// TIA Portal project "Robotino" (V18)

(* hardware
DEVICE "S7-1500/ET200MP-Station_1"  S7-1500 station
   slot 0: "Profilschiene_0"  Rack  6ES7 590-1***0-0AA0
   slot 1: "PLC_1"  CPU 1516-3 PN/DP  6ES7 516-3AP03-0AB0  V3.0
      slot 3: "CPU-Display_1"  6ES7591-1BA00-0AA0
      slot 32768: "PROFINET-Schnittstelle_1"  X1
      slot 33024: "PROFINET-Schnittstelle_2"  X2
      slot 33280: "DP-Schnittstelle_1"  X3
      slot 34817: "Virtual CP interface port_1"  Virtual CP interface port  Virtual CP interface port
   slot 2: "DI 32x24VDC HF_1"  DI 32x24VDC HF  6ES7 521-1BL00-0AB0  V2.2
   slot 3: "DQ 32x24VDC/0.5A HF_1"  DQ 32x24VDC/0.5A HF  6ES7 522-1BL01-0AB0  V1.1
   slot 4: "AI 8xU/I/RTD/TC ST_1"  AI 8xU/I/RTD/TC ST  6ES7 531-7KF00-0AB0  V2.2
   slot 5: "AQ 4xU/I ST_1"  AQ 4xU/I ST  6ES7 532-5HD00-0AB0  V2.2
DEVICE "ROBOTINO_HMI"  MTP700 Unified Comfort
   slot 0: "ROBOTINO_HMI"  MTP700 Unified Comfort  6AV2 128-3GB06-0AXx  18.0.0.2
   slot 1: "HMI_RT_1"  MTP700 Unified Comfort  6AV2 128-3GB06-0AXx  18.0.0.2
   slot 5: "ROBOTINO_HMI.IE_CP_1"  PROFINET Interface  18.0.0.2
      slot 1: "PROFINET Schnittstelle_1"  PROFINET Interface
         slot 1: "Port_1"  Port
         slot 2: "Port_2"  Port
   slot 6: "ROBOTINO_HMI.IE_CP_2"  PROFINET Interface  18.0.0.2
      slot 1: "PROFINET Schnittstelle_GBit"  PROFINET Interface
         slot 1: "Port_1"  Port
*)

// ===== PLC "PLC_1"  CPU 1516-3 PN/DP =====

DATA_BLOCK "OPCUA"   // DB1
{ S7_Optimized_Access := 'TRUE' }
VERSION : 0.1
   VAR
      Test_bool : Bool;
      Test_int : Int;
      Test_String : String;
      Test_array_bool : Array[0..1] of Bool;
      Test_array_int : Array[0..1] of Int;
   END_VAR
BEGIN
END_DATA_BLOCK

DATA_BLOCK "ROBOTINO"   // DB2
{ S7_Optimized_Access := 'TRUE' }
VERSION : 0.1
   VAR
      Bumper : Bool;
      Distance_Sensors : Array[1..9] of Real;
      Digital_Inputs : Array[1..8] of Bool;
      Analog_Inputs : Array[1..8] of Real;
      Motor4 : Int;   // Belt
      Motor4_Current : Real;
      Digital_Outputs : Array[1..8] of Bool;
      Digital_Outputs_Status : Array[1..8] of Bool;
      Relay : Array[1..2] of Bool;
      Relay_Status : Array[1..2] of Bool;
      Odometry : Array[0..6] of Real;
      Omnidrive : Array[0..2] of Real;
      Bat_Voltage : Real;
      Charging_State : String;
      Charging_Current : Real;
      Controller_Info : Array[0..1] of String;
      Image_Version : String;
      Factory_Status : Array[0..3] of Bool;
      Position_ID : Int;
      Start_GoToPos : Bool;
      GoToPos_Completed : Bool;
      Robotino_Position : Int;   // actual defined position of robotino. =0 If robotino is not on a defined position
      DockTo_Completed : Bool;   // =1 if robotino is docked
      Start_DockTo : Bool;
      Stop_DockTo : Bool;
   END_VAR
BEGIN
   // Digital_Inputs[3] : Vision Sensor Package Present
   // Digital_Inputs[4] : IR Station Ready (false connected)
   // Digital_Inputs[5] : Reset Button
   // Digital_Outputs[3] : lamp tower red
   // Digital_Outputs[4] : lamp tower yellow
   // Digital_Outputs[5] : lamp tower green
   // Digital_Outputs[6] : light reset button
   // Digital_Outputs[1] : IR Robotino Ready
   // Digital_Outputs_Status[1] : IR Robotino Ready
   // Digital_Outputs_Status[3] : lamp tower red
   // Digital_Outputs_Status[4] : lamp tower yellow
   // Digital_Outputs_Status[5] : lamp tower green
   // Digital_Outputs_Status[6] : light reset button
   // Relay_Status[1] : Enable analog sensors
   // Odometry[0] : x /m
   // Odometry[1] : y /m
   // Odometry[2] : rot /rad
   // Odometry[3] : vx
   // Odometry[4] : vy
   // Odometry[5] : omega
   // Odometry[6] : sequence number
   // Omnidrive[0] : vx
   // Omnidrive[1] : vy
   // Omnidrive[2] : omega
   // Relay[1] : Enable analog sensors
   // Analog_Inputs[1] : Distance Left (not scaled)
   // Analog_Inputs[2] : Distance Center (not scaled)
   // Analog_Inputs[3] : Distance Right (not scaled)
   // Controller_Info[1] : Software version
   // Controller_Info[0] : Hardware version
   // Factory_Status[0] : Idle
   // Factory_Status[1] : Busy
   // Factory_Status[2] : Error
   // Factory_Status[3] : Started
   // Digital_Inputs[1] : Emergncy Button
END_DATA_BLOCK

DATA_BLOCK "GoTo_DB"   // DB3
{ S7_Optimized_Access := 'TRUE' }
VERSION : 0.1
// stored: InstanceOfName GoTo
"GoTo"
BEGIN
END_DATA_BLOCK

DATA_BLOCK "DockTo_DB"   // DB5
{ S7_Optimized_Access := 'TRUE' }
VERSION : 0.1
// stored: InstanceOfName DockTo
"DockTo"
BEGIN
END_DATA_BLOCK

DATA_BLOCK "Robotino_Control"   // DB6
{ S7_Optimized_Access := 'TRUE' }
VERSION : 0.1
   VAR
      Start_GoTo : Bool;
      Start_DockTo : Bool;
      Ready_DockTo : Bool;
      Stop_DockTo : Bool;
      Conveyor : Int;
      PosId : Int;
   END_VAR
BEGIN
END_DATA_BLOCK

// folder: System blocks/Program resources

DATA_BLOCK "IEC_Timer_0_DB"   // DB4
{ S7_Optimized_Access := 'TRUE' }
AUTHOR : Simatic
FAMILY : IEC
NAME : IEC_TMR
VERSION : 1.0
// stored: InstanceOfName IEC_TIMER
"IEC_TIMER"
BEGIN
END_DATA_BLOCK

DATA_BLOCK "IEC_Timer_0_DB_1"   // DB8
{ S7_Optimized_Access := 'TRUE' }
AUTHOR : Simatic
FAMILY : IEC
NAME : IEC_TMR
VERSION : 1.0
// stored: InstanceOfName IEC_TIMER
"IEC_TIMER"
BEGIN
END_DATA_BLOCK

// folder: (top level)

FUNCTION_BLOCK "GoTo"   // FB1, FBD
{ S7_Optimized_Access := 'TRUE' }
VERSION : 0.1
   VAR_INPUT
      Idle : Bool;
      Busy : Bool;
      Error : Bool;
      Started : Bool;
      Pos : Int;
      Start : Bool;
   END_VAR
   VAR_OUTPUT
      GoTo_Completed : Bool;
      GoTo_Start : Bool;
      GoTo_PosId : Int;
      actual_PosId : Int;
   END_VAR
   VAR_TEMP
      process_completed : Bool;
      busy_negedge : Bool;
      idle_posedge : Bool;
      process_started : Bool;
      completed_p_edge : Bool;
   END_VAR
   VAR_TEMP   // added for the SCL form of the ladder/FBD networks
      _w1 : Bool;
   END_VAR
BEGIN

REGION Network 1
   // Anzahl definierter Positionen in Factory ggf. anpassen
   // 
   // Sinnhaftigkeit von TOF und Zeit prüfen
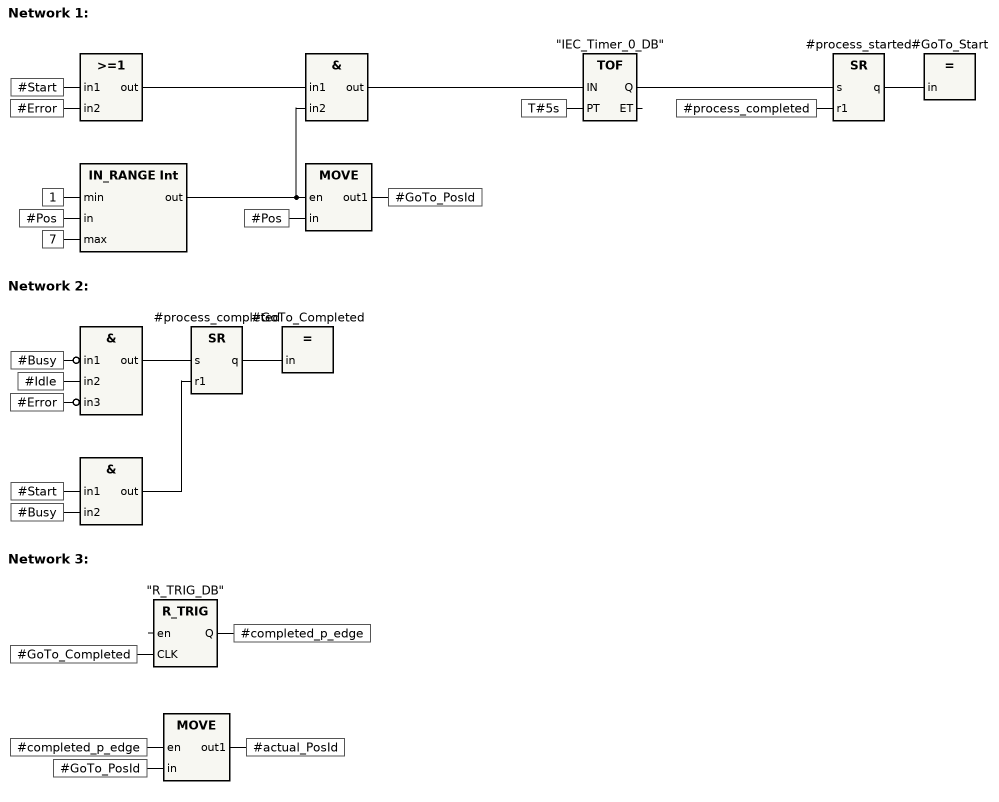
   #_w1 := (1 <= #Pos) AND (#Pos <= 7);
   "IEC_Timer_0_DB".TOF(IN := (#Start OR #Error) AND #_w1, PT := T#5s);
   IF "IEC_Timer_0_DB".Q THEN
       #process_started := TRUE;   // SR flip-flop
   END_IF;
   IF #process_completed THEN #process_started := FALSE; END_IF;
   #GoTo_Start := #process_started;
   IF #_w1 THEN #GoTo_PosId := #Pos; END_IF;
END_REGION

REGION Network 2
   // Startbefehl nach GoToCompleted zurückssetzen
   IF NOT #Busy AND #Idle AND NOT #Error THEN
       #process_completed := TRUE;   // SR flip-flop
   END_IF;
   IF #Start AND #Busy THEN #process_completed := FALSE; END_IF;
   #GoTo_Completed := #process_completed;
END_REGION

REGION Network 3
   // Registrierung der aktuellen Position
   // nur p edge als enable nehemen
   "R_TRIG_DB"(CLK := #GoTo_Completed, Q => #completed_p_edge);   // R_TRIG
   IF #completed_p_edge THEN #actual_PosId := #GoTo_PosId; END_IF;
END_REGION
END_FUNCTION_BLOCK

FUNCTION_BLOCK "DockTo"   // FB2, GRAPH_PLUS
{ S7_Optimized_Access := 'TRUE' }
VERSION : 0.1
   VAR_INPUT
      OFF_SQ : Bool := false;
      INIT_SQ : Bool := false;
      ACK_EF : Bool := false;
      S_PREV : Bool := false;
      S_NEXT : Bool := false;
      SW_AUTO : Bool := false;
      SW_TAP : Bool := false;
      SW_TOP : Bool := false;
      SW_MAN : Bool := false;
      S_SEL : Int := 0;
      S_ON : Bool := false;
      S_OFF : Bool := false;
      T_PUSH : Bool := false;
      idle : Bool;
      busy : Bool;
      error_factory : Bool;
      robotino_position : Int;
      distance_left : Real;
      distance_center : Real;
      distance_right : Real;
   END_VAR
   VAR_OUTPUT
      S_NO : Int := 0;
      S_MORE : Bool := false;
      S_ACTIVE : Bool := false;
      ERR_FLT : Bool := false;
      AUTO_ON : Bool := false;
      TAP_ON : Bool := false;
      TOP_ON : Bool := false;
      MAN_ON : Bool := false;
      docking_completed : Bool;
      docking_started : Bool;
      vx : Real;
      vy : Real;
      omega : Real;
      relay_analogsensors : Bool;
   END_VAR
   VAR
      HMI_INFO : Array[0..8] of UInt;
      IF_PAR : G7_IfParPlus_V6;
      RT_DATA : G7_RTDataPlus_V6;
      Trans1 : G7_TransitionPlus_V6;
      Trans2 : G7_TransitionPlus_V6;
      Trans3 : G7_TransitionPlus_V6;
      Trans4 : G7_TransitionPlus_V6;
      Trans5 : G7_TransitionPlus_V6;
      Trans6 : G7_TransitionPlus_V6;
      Trans7 : G7_TransitionPlus_V6;
      Trans8 : G7_TransitionPlus_V6;   // Transitionsstruktur
      Trans9 : G7_TransitionPlus_V6;   // Transitionsstruktur
      Trans10 : G7_TransitionPlus_V6;   // Transitionsstruktur
      Trans11 : G7_TransitionPlus_V6;   // Transitionsstruktur
      Trans13 : G7_TransitionPlus_V6;   // Transitionsstruktur
      Trans14 : G7_TransitionPlus_V6;   // Transitionsstruktur
      Trans18 : G7_TransitionPlus_V6;   // Transitionsstruktur
      Step1 : G7_StepPlus_V6;
      Step2 : G7_StepPlus_V6;
      Step3 : G7_StepPlus_V6;
      Step4 : G7_StepPlus_V6;
      Step5 : G7_StepPlus_V6;
      Step6 : G7_StepPlus_V6;
      Step7 : G7_StepPlus_V6;   // Schrittstruktur
      Step8 : G7_StepPlus_V6;   // Schrittstruktur
      Step9 : G7_StepPlus_V6;   // Schrittstruktur
      Step11 : G7_StepPlus_V6;   // Schrittstruktur
      Step13 : G7_StepPlus_V6;   // Schrittstruktur
      Step14 : G7_StepPlus_V6;   // Schrittstruktur
      SINI : Array[0..1] of USInt;
      LSTT : Array[0..13] of USInt;
      ATAJ : Array[0..13] of USInt;
      ATAB : Array[0..13] of USInt;
      PSTT : Array[0..13] of USInt;
      NSTT : Array[0..13] of USInt;
      ASSJ : Array[0..11] of USInt;
      ASSB : Array[0..11] of USInt;
      PTTS : Array[0..11] of USInt;
      NTTS : Array[0..11] of USInt;
      SW_SQTS : Array[0..11] of USInt;
      SWITCH : Array[0..6] of USInt;
      TVX : Array[0..5] of USInt;
      TTX : Array[0..5] of USInt;
      TSX : Array[0..1] of USInt;
      S00X : Array[0..1] of USInt;
      SOFFX : Array[0..1] of USInt;
      SONX : Array[0..1] of USInt;
      SAX : Array[0..1] of USInt;
      SERRX : Array[0..12] of USInt;
      SMX : Array[0..12] of USInt;
      S0X : Array[0..12] of USInt;
      S1X : Array[0..12] of USInt;
      IL_ALARM_INST : Diag_Alarm;
      SUP_ALARM_INST : Diag_Alarm;
      STEP_TIME_ALARM_INST : Diag_Alarm;
      IEC_TIMER_INST : IEC_TIMER;
      TRANSACTION_FLAG : Bool := false;
   END_VAR
   VAR CONSTANT
      threshold_x : Real := 1.5;
      threshold_y : Real := 1.4;
   END_VAR
   // SINI[0] := 2;
   // LSTT[0] := 255;
   // ATAJ[1] := 1;
   // ATAB[1] := 1;
   // PSTT[1] := 1;
   // NSTT[0] := 3;
   // ASSJ[1] := 1;
   // ASSB[1] := 1;
   // PTTS[0] := 255;
   // NTTS[1] := 1;
   // TVX[0] := 16#1;
   // TTX[0] := 16#1;
   // TSX[0] := 16#1;
   // S00X[0] := 16#1;
   // SOFFX[0] := 16#1;
   // SONX[0] := 16#1;
   // SAX[0] := 16#1;
   // SERRX[0] := 16#1;
   // SMX[0] := 16#1;
   // S0X[0] := 16#1;
   // S1X[0] := 16#1;
   // LSTT[1] := 255;
   // ATAJ[2] := 2;
   // ATAB[2] := 2;
   // PSTT[2] := 2;
   // NSTT[1] := 6;
   // ASSJ[2] := 2;
   // ASSB[2] := 2;
   // PTTS[2] := 9;
   // NTTS[2] := 2;
   // LSTT[3] := 255;
   // LSTT[4] := 255;
   // LSTT[5] := 255;
   // LSTT[6] := 255;
   // ATAJ[3] := 3;
   // ATAJ[4] := 4;
   // ATAJ[5] := 5;
   // ATAJ[6] := 6;
   // ATAB[3] := 4;
   // ATAB[4] := 3;
   // ATAB[5] := 5;
   // ATAB[6] := 6;
   // PSTT[3] := 3;
   // PSTT[4] := 3;
   // PSTT[5] := 5;
   // PSTT[6] := 4;
   // NSTT[3] := 5;
   // NSTT[4] := 4;
   // NSTT[5] := 1;
   // NSTT[6] := 10;
   // ASSJ[3] := 3;
   // ASSJ[4] := 4;
   // ASSJ[5] := 5;
   // ASSB[3] := 3;
   // ASSB[4] := 4;
   // ASSB[5] := 5;
   // PTTS[1] := 5;
   // PTTS[4] := 4;
   // PTTS[5] := 3;
   // NTTS[3] := 3;
   // NTTS[4] := 6;
   // NTTS[5] := 5;
   // SW_SQTS[1] := 1;
   // SW_SQTS[2] := 2;
   // SW_SQTS[4] := 3;
   // SW_SQTS[5] := 1;
   // LSTT[7] := 255;
   // ATAJ[7] := 7;
   // ATAB[7] := 8;
   // PSTT[7] := 9;
   // NSTT[7] := 7;
   // ASSJ[6] := 6;
   // ASSB[6] := 6;
   // PTTS[6] := 1;
   // NTTS[6] := 11;
   // SW_SQTS[6] := 1;
   // LSTT[8] := 255;
   // LSTT[9] := 255;
   // LSTT[10] := 255;
   // ATAJ[8] := 8;
   // ATAJ[9] := 10;
   // ATAJ[10] := 9;
   // ATAB[8] := 7;
   // ATAB[9] := 9;
   // ATAB[10] := 10;
   // PSTT[8] := 9;
   // PSTT[9] := 7;
   // PSTT[10] := 8;
   // NSTT[8] := 8;
   // NSTT[9] := 2;
   // NSTT[10] := 2;
   // ASSJ[7] := 7;
   // ASSJ[8] := 8;
   // ASSB[7] := 7;
   // ASSB[8] := 8;
   // PTTS[7] := 7;
   // PTTS[8] := 8;
   // NTTS[7] := 9;
   // NTTS[8] := 10;
   // SW_SQTS[7] := 4;
   // SW_SQTS[8] := 5;
   // LSTT[11] := 255;
   // LSTT[12] := 255;
   // LSTT[13] := 255;
   // ATAJ[11] := 13;
   // ATAJ[12] := 12;
   // ATAJ[13] := 11;
   // ATAB[11] := 11;
   // ATAB[12] := 12;
   // ATAB[13] := 13;
   // PSTT[11] := 6;
   // PSTT[12] := 10;
   // PSTT[13] := 11;
   // NSTT[11] := 9;
   // NSTT[12] := 11;
   // NSTT[13] := 9;
   // ASSJ[9] := 9;
   // ASSJ[10] := 10;
   // ASSJ[11] := 11;
   // ASSB[9] := 9;
   // ASSB[10] := 10;
   // ASSB[11] := 11;
   // PTTS[9] := 11;
   // PTTS[10] := 6;
   // PTTS[11] := 12;
   // NTTS[9] := 7;
   // NTTS[10] := 12;
   // NTTS[11] := 13;
   // SW_SQTS[9] := 6;
   // SW_SQTS[10] := 3;
   // SW_SQTS[11] := 3;
BEGIN
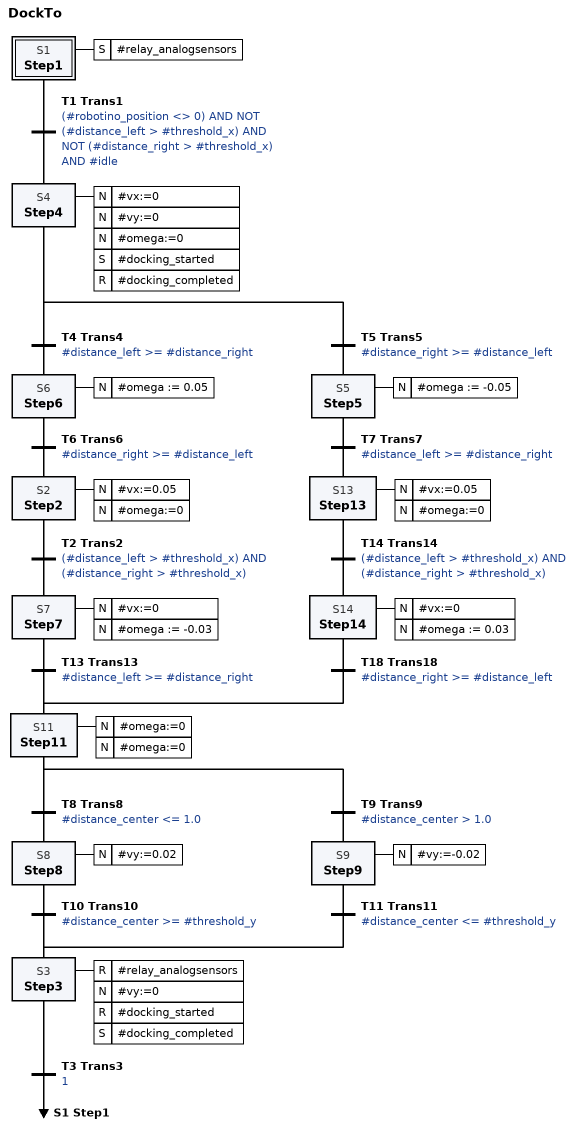
   // sequencer 1
   INITIAL_STEP Step1:   // S1, max time T#10S, warning time T#7S
              S    #relay_analogsensors
   END_STEP
   TRANSITION Trans1 FROM Step1 TO Step4   // T1
      := (#robotino_position <> 0) AND NOT (#distance_left > #threshold_x) AND NOT (#distance_right > #threshold_x) AND #idle;
   END_TRANSITION
   STEP Step2:   // S2, max time T#10S, warning time T#7S
              N    #vx:=0.05
              N    #omega:=0
   END_STEP
   TRANSITION Trans2 FROM Step2 TO Step7   // T2
      := (#distance_left > #threshold_x) AND (#distance_right > #threshold_x);
   END_TRANSITION
   STEP Step3:   // S3, max time T#10S, warning time T#7S
              R    #relay_analogsensors
              N    #vy:=0
              R    #docking_started
              S    #docking_completed
   END_STEP
   TRANSITION Trans3 FROM Step3 TO Step1   // T3, jump
      := 1;
   END_TRANSITION
   STEP Step4:   // S4, max time T#10S, warning time T#7S
              N    #vx:=0
              N    #vy:=0
              N    #omega:=0
              S    #docking_started
              R    #docking_completed
   END_STEP
   TRANSITION Trans4 FROM Step4 TO Step6   // T4
      := #distance_left >= #distance_right;
   END_TRANSITION
   TRANSITION Trans5 FROM Step4 TO Step5   // T5
      := #distance_right >= #distance_left;
   END_TRANSITION
   STEP Step5:   // S5, max time T#10S, warning time T#7S
              N    #omega := -0.05
   END_STEP
   TRANSITION Trans7 FROM Step5 TO Step13   // T7
      := #distance_left >= #distance_right;
   END_TRANSITION
   STEP Step6:   // S6, max time T#10S, warning time T#7S
              N    #omega := 0.05
   END_STEP
   TRANSITION Trans6 FROM Step6 TO Step2   // T6
      := #distance_right >= #distance_left;
   END_TRANSITION
   STEP Step7:   // S7, max time T#10S, warning time T#7S
              N    #vx:=0
              N    #omega := -0.03
   END_STEP
   TRANSITION Trans13 FROM Step7 TO Step11   // T13
      := #distance_left >= #distance_right;
   END_TRANSITION
   STEP Step8:   // S8, max time T#10S, warning time T#7S
              N    #vy:=0.02
   END_STEP
   TRANSITION Trans10 FROM Step8 TO Step3   // T10
      := #distance_center >= #threshold_y;
   END_TRANSITION
   STEP Step9:   // S9, max time T#10S, warning time T#7S
              N    #vy:=-0.02
   END_STEP
   TRANSITION Trans11 FROM Step9 TO Step3   // T11
      := #distance_center <= #threshold_y;
   END_TRANSITION
   STEP Step11:   // S11, max time T#10S, warning time T#7S
              N    #omega:=0
              N    #omega:=0
   END_STEP
   TRANSITION Trans8 FROM Step11 TO Step8   // T8
      := #distance_center <= 1.0;
   END_TRANSITION
   TRANSITION Trans9 FROM Step11 TO Step9   // T9
      := #distance_center > 1.0;
   END_TRANSITION
   STEP Step13:   // S13, max time T#10S, warning time T#7S
              N    #vx:=0.05
              N    #omega:=0
   END_STEP
   TRANSITION Trans14 FROM Step13 TO Step14   // T14
      := (#distance_left > #threshold_x) AND (#distance_right > #threshold_x);
   END_TRANSITION
   STEP Step14:   // S14, max time T#10S, warning time T#7S
              N    #vx:=0
              N    #omega := 0.03
   END_STEP
   TRANSITION Trans18 FROM Step14 TO Step11   // T18
      := #distance_right >= #distance_left;
   END_TRANSITION
END_FUNCTION_BLOCK

ORGANIZATION_BLOCK "Main"   // OB1, FBD, ProgramCycle
{ S7_Optimized_Access := 'TRUE' }
VERSION : 0.1
   VAR_INPUT
      Initial_Call : Bool;
      Remanence : Bool;
   END_VAR
BEGIN

REGION Network 1: HMI
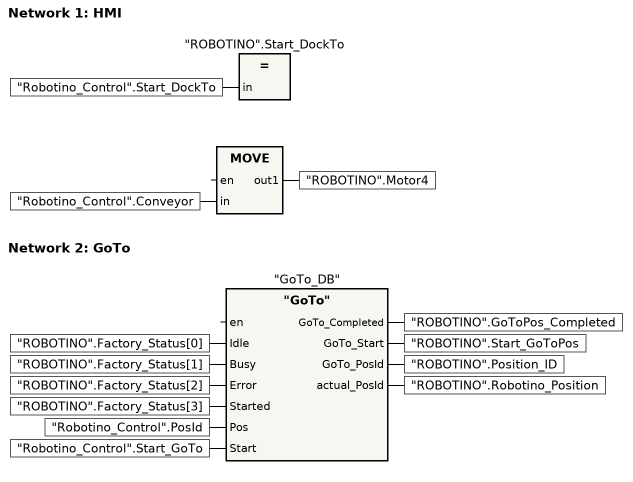
   "ROBOTINO".Start_DockTo := "Robotino_Control".Start_DockTo;
   "ROBOTINO".Motor4 := "Robotino_Control".Conveyor;
END_REGION

REGION Network 2: GoTo
   "GoTo_DB"(Idle := "ROBOTINO".Factory_Status[0],   // "GoTo"
             Busy := "ROBOTINO".Factory_Status[1],
             Error := "ROBOTINO".Factory_Status[2],
             Started := "ROBOTINO".Factory_Status[3],
             Pos := "Robotino_Control".PosId,
             Start := "Robotino_Control".Start_GoTo,
             GoTo_Completed => "ROBOTINO".GoToPos_Completed,
             GoTo_Start => "ROBOTINO".Start_GoToPos,
             GoTo_PosId => "ROBOTINO".Position_ID,
             actual_PosId => "ROBOTINO".Robotino_Position);
END_REGION

REGION Network 3: DockTo
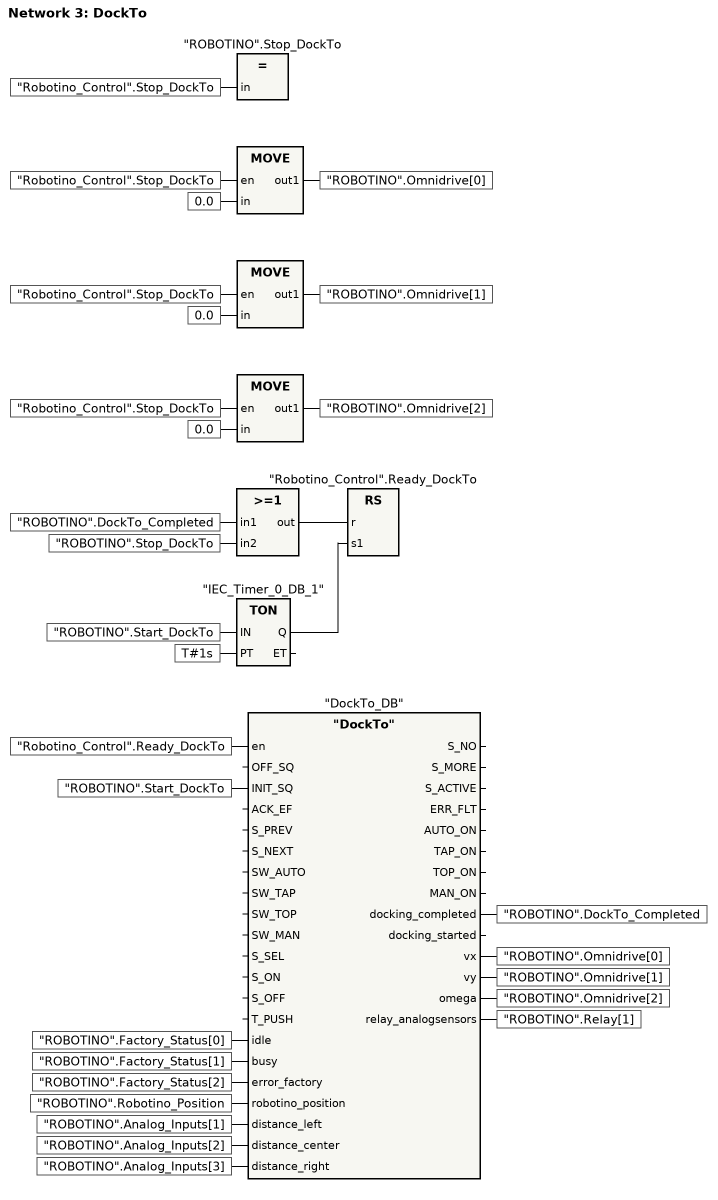
   "ROBOTINO".Stop_DockTo := "Robotino_Control".Stop_DockTo;
   IF "Robotino_Control".Stop_DockTo THEN
       "ROBOTINO".Omnidrive[0] := 0.0;
       "ROBOTINO".Omnidrive[1] := 0.0;
       "ROBOTINO".Omnidrive[2] := 0.0;
   END_IF;
   "IEC_Timer_0_DB_1".TON(IN := "ROBOTINO".Start_DockTo, PT := T#1s);
   IF "ROBOTINO".DockTo_Completed OR "ROBOTINO".Stop_DockTo THEN
       "Robotino_Control".Ready_DockTo := FALSE;   // RS flip-flop
   END_IF;
   IF "IEC_Timer_0_DB_1".Q THEN "Robotino_Control".Ready_DockTo := TRUE; END_IF;
   IF "Robotino_Control".Ready_DockTo THEN
       "DockTo_DB"(INIT_SQ := "ROBOTINO".Start_DockTo,   // "DockTo"
                   idle := "ROBOTINO".Factory_Status[0],
                   busy := "ROBOTINO".Factory_Status[1],
                   error_factory := "ROBOTINO".Factory_Status[2],
                   robotino_position := "ROBOTINO".Robotino_Position,
                   distance_left := "ROBOTINO".Analog_Inputs[1],
                   distance_center := "ROBOTINO".Analog_Inputs[2],
                   distance_right := "ROBOTINO".Analog_Inputs[3],
                   docking_completed => "ROBOTINO".DockTo_Completed,
                   vx => "ROBOTINO".Omnidrive[0],
                   vy => "ROBOTINO".Omnidrive[1],
                   omega => "ROBOTINO".Omnidrive[2],
                   relay_analogsensors => "ROBOTINO".Relay[1]);
   END_IF;
END_REGION
END_ORGANIZATION_BLOCK

(* ===== HMI "HMI_RT_1" =====
connection "HMI_Verbindung_1": ETHERNET, ILRT_S7_1500_OMS

HMI tags "Standard-Variablentabelle"
   "Robotino_Control_Start_GoTo" : Bool = PLC Robotino_Control.Start_GoTo, T100ms
   "Robotino_Control_Start_DockTo" : Bool = PLC Robotino_Control.Start_DockTo, T100ms
   "Robotino_Control_Stop_DockTo" : Bool = PLC Robotino_Control.Stop_DockTo, T100ms
   "Robotino_Control_Conveyor" : Int = PLC Robotino_Control.Conveyor, T100ms
   "Robotino_Control_PosId" : Int = PLC Robotino_Control.PosId, T100ms
   "ROBOTINO_Digital_Inputs{1}" : Bool = PLC ROBOTINO.Digital_Inputs[1] AT %DB1.DBW0, T100ms
   "ROBOTINO_Digital_Outputs_Status{3}" : Bool = PLC ROBOTINO.Digital_Outputs_Status[3], T100ms
   "ROBOTINO_Digital_Outputs_Status{4}" : Bool = PLC ROBOTINO.Digital_Outputs_Status[4], T100ms
   "ROBOTINO_Digital_Outputs_Status{5}" : Bool = PLC ROBOTINO.Digital_Outputs_Status[5], T100ms

text list "SystemTextList_ConfigErrorAlarmTextLibrary_1": 1 'NameService Konfigurationsfehler: Implizites Löschen. Subelement-Instanz @6%s@ muss explizit gelöscht werden.'; 2 'NameService Konfigurationsfehler: Implizites Löschen. Alias/Format/Unit-Instanz @6%s@ muss explizit gelöscht werden.'

text list "SystemTextList_ConfigErrorAlarmTextLibrary_2": 1 'EvDpManager::cleanupDeletedDatapoint - alert handler config is deleted implicitly for deleted datapoint, @3%s@'; 2 'EvDpManager::cleanupDeletedDatapoint - alert handler config is deleted implicitly but still has overrides, @3%s@'; 3 'EvDpManager::cleanupDeletedDatapoint - default value config is deleted implicitly for deleted datapoint, @3%s@'; 4 'EvDpManager::cleanupDeletedDatapoint - default value config is deleted implicitly but still has overrides, @3%s@'; 5 'EvDpManager::cleanupDeletedDatapoint - initial value config is deleted implicitly for deleted datapoint, @3%s@'; 6 'EvDpManager::cleanupDeletedDatapoint - initial value config is deleted implicitly but still has overrides, @3%s@'; 7 'EvDpManager::cleanupDeletedDatapoint - distribution config is deleted implicitly for deleted datapoint, @3%s@'; 8 'EvDpManager::cleanupDeletedDatapoint - distribution config is deleted implicitly but still has overrides, @3%s@'; 9 'EvDpManager::cleanupDeletedDatapoint - rangeCheck config is deleted implicitly for deleted datapoint, @3%s@'; 10 'EvDpManager::cleanupDeletedDatapoint - rangeCheck config is deleted implicitly but still has overrides, @3%s@'

text list "SystemTextList_ConfigErrorAlarmTextLibrary_3": 1 'Der konfigurierte Datenpunkttyp wurde gelöscht. Ein konfigurierter Typ ist aber noch für den Knotentyp definiert: @3%s@.'; 2 'Der konfigurierter Datenpunkt-Knotentyp wurde im Datenpunkttyp gelöscht. Ein konfigurierter Typ ist aber noch für das Element definiert: @3%s@.'

text list "SystemTextList_ConfigErrorAlarmTextLibrary_4": 2 'Zyklen: @6%s@ existiert nicht'; 3 'Alarme: @6%s@ existiert bereits'; 4 'Variablen: Adresse @6%s@ wurde abgelehnt'; 1 'Verbindungen: @6%s@ existiert nicht'; 5 'Variablen: Erfassungsart @6%s@ wird nicht unterstützt.'; 6 'Zyklen: @6%s@ wurde gelöscht aber zugehörige Variablen existieren.'; 7 'Verbindungen: @6%s@ wurde gelöscht aber zugehörige Variablen existieren.'; 8 'Variablen: Variable @6%s@ wurde abgelehnt.'; 9 'Variablen: Variable @6%s@ hat einen ungültigen Wert.'; 0 'Verbindungen: Verbindung zu @6%s@ konnte nicht hergestellt werden.'; 65638 'Verbindungen: Verbindung zu @6%s@ konnte nicht hergestellt werden.'; 65639 'Verbindungen: @6%s@ getrennt.'; 65640 'Verbindungen: Verbindung zum HMI-Gerät @6%s@ getrennt.'; 65641 'Verbindungen: Verbindung zur PLC @6%s@ getrennt.'; 65541 'Verbindungen: Zeitüberschreitung beim Aufbau der Verbindung zu @6%s@.'; 65542 'Verbindungen: @6%s@ gestört.'; 65543 'Verbindungen: Verbindung zum HMI-Gerät getrennt. Verbindung @5%s@ wurde geändert.'; 65544 'Verbindungen: Verbindung zum HMI-Gerät getrennt. Treibereigenschaft wurde geändert bei Verbindung @5%s@.'

text list "SystemTextList_ConfigErrorAlarmTextLibrary_5": 1 'Verbindungen: Zyklus der Lebenszeichenüberwachung muss kleiner sein als die Antwortzeit.'; 2 'Verbindungen: Zyklische Dienste sind konfiguriert, werden aber vom Zielgerät nicht unterstützt.'; 3 'Verbindungen: Änderungsgesteuertes Lesen ist konfiguriert, wird aber vom Zielgerät nicht unterstützt.'; 4 'Variablen: Die Adresse @6%s@ existiert in der PLC nicht.'; 5 'Variablen: Der Standardkonvertierungstyp für die Adresse @6%s@ konnte nicht ermittelt werden.'; 6 'Variablen: Ungültiger Konvertierungstyp'; 7 'Zyklen: Ungültiger Konvertierungstyp. Konvertierung wird nicht unterstützt am HmiCycle.'; 4096 'Verbindungen: Version der Adresse @6%s@ wird nicht unterstützt.'; 4097 'Verbindungen: Profibus-Adresse wird nicht unterstützt.'; 4098 'Verbindungen: Softbus-Adresse wird nicht unterstützt.'; 4099 'Verbindungen: Adressetyp @6%s@ wird nicht unterstützt.'; 4100 'Verbindungen: Ungültiger Verbindungsname @6%s@. Zugriffspunkt wird ignoriert.'; 4101 'Verbindungen: Routing wird nicht unterstützt. @6%s@ wird nicht verwendet.'; 4102 'Verbindungen: Routing werden nicht unterstützt. @6%s@ wird nicht verwendet.'; 4103 'Verbindungen: Ungültige IP-Adresse @6%s@'; 4104 'Verbindungen: Ungültige Named Connection @6%s@. Gültiges Format: >VMD</>Verbindung<'; 4105 'Verbindungen: Ungültige Named Connection @6%s@. VMD Verbindungsname ist zu lang. Es sind nur 24 Zeichen erlaubt.'; 4106 'Verbindungen: Ungültige Named Connection @6%s@. Verbindungsname ist zu lang. Es sind nur 32 Zeichen erlaubt.'; 4107 'Verbindungen: Rack-Nummer @6%s@ ist außerhalb des erlaubten Bereichs (0..7)'; 4108 'Verbindungen: Ungültige Named Connection @6%s@. Rack wird ignoriert.'; 4109 'Verbindungen: Slot-Nummer @6%s@ ist außerhalb des erlaubten Bereichs (1..32)'; 4110 'Verbindungen: Ungültige Named Connection @6%s@. Slot wird ignoriert.'; 4111 'Verbindung konnte nicht hergestellt werden. Maximale Anzahl von verfügbaren Verbindungen (@6%s@) ist überschritten.'; 4112 'Verbindung abgebrochen. Kein Lebenszeichen in den letzten @4%s@ ms.'; 4113 'Verbindung konnte nicht hergestellt werden - @4%s@'; 4114 'Verbindung konnte nicht hergestellt werden. Die Adresse @6%s@ kann nicht verwendet werden.'; 4115 'Verbindung konnte nicht hergestellt werden. Ungültige Adresse @6%s@'; 4116 'Verbindung konnte nicht hergestellt werden - @4%s@'

text list "SystemTextList_ConfigErrorAlarmTextLibrary_6": 1 'Verbindung konnte nicht hergestellt werden. Applikation-Instanz-Zertifikat ist nicht konfiguriert.'; 2 'Verbindung konnte nicht hergestellt werden. Server hat das Client-Zertifikat abgelehnt. OPC UA Status Code @4%s@.'; 3 'Verbindung konnte nicht hergestellt werden. Internes Problem im Zertifikatspeicher. OPC UA Status Code @4%s@'; 4 'Verbindung konnte nicht hergestellt werden. Applikation-Instanz-Zertifikat konnte nicht geladen werden. OPC UA Status Code @5%s@'; 5 'Verbindung konnte nicht hergestellt werden. Server hat kein Zertifikat zur Verfügung gestellt. @4%s@'; 6 'Verbindung konnte nicht hergestellt werden. Validierung vom Server-Zertifikat ist fehlgeschlagen. OPC UA Status Code @4%s@.'; 7 'Verbindung wurde geschlossen. Fehler bei der Alarmsynchronisation. OPC UA Status Code @4%s@.'; 8 'Verbindung wurde geschlossen. Alarm/Event Subscription ist fehlgeschlagen. Die Anzahl der Operationen auf dem Server wurde überschritten.'; 9 'Verbindung wurde geschlossen. Alarm/Event Subscription ist fehlgeschlagen. Die Anzahl der Alarm/Event Subscriptions auf dem Server wurde überschritten.'; 10 'Verbindung konnte nicht hergestellt werden. Server meldet ein Lizenzproblem. OPC UA Status Code @4%s@.'; 11 'Verbindung konnte nicht hergestellt werden. Maximale Anzahl an Server-Sitzungen wurde überschritten.'; 12 'Verbindung konnte nicht hergestellt werden. Sicherheitskonfiguration ist inkonsistent. @4%s@'; 13 'Verbindung konnte nicht hergestellt werden. Die Adresse @4%s@ kann nicht verwendet werden.'; 14 'Verbindung konnte nicht hergestellt werden. OPC UA Status Code @4%s@'; 15 'Verbindung abgebrochen. OPC UA Server wurde gestoppt.'; 16 'Verbindung abgebrochen. Kein Lebenszeichen in den letzten @4%s@ ms.'; 17 'Verbindung wurde geschlossen - OPC UA Server-Wartung.'; 18 'Verbindung konnte nicht hergestellt werden. Ungültige Konfiguration des Authentifizierungsmodus - @4%s@'; 19 'Verbindung konnte nicht hergestellt werden. Anwender konnte nicht authentifiziert werden. OPC UA Status Code @4%s@'; 20 'Verbindung konnte nicht hergestellt werden. Server erlaubt keine anonyme Verbindung. OPC UA Status Code @4%s@'; 21 'Verbindung konnte nicht hergestellt werden. Zertifikatsproblem: Fehler beim Schreiben der sicherheitsrelevanten Daten nach @4%s@.'; 22 'Verbindung konnte nicht hergestellt werden. Zertifikatsproblem: Unerwartete Datei im Verzeichnis @4%s@ kann nicht entfernt werden.'; 23 'Verbindung konnte nicht hergestellt werden. Benutzer konnte nicht authentifiziert werden. Kein Benutzer oder Passwort konfiguriert.'; 24 'Verbindung konnte nicht hergestellt werden. Unerwartete Länge vom Server-Zertifikat. @4%s@'; 25 'Verbindung konnte nicht hergestellt werden. @4%s@ ohne Inhalt.'; 26 'Verbindung konnte nicht hergestellt werden. @4%s@ hat ein unerwartetes Format.'; 27 'Verbindung konnte nicht hergestellt werden. Server-Endpunkte können nicht gelesen werden. OPC UA Status Code @4%s@'; 28 'Verbindung konnte nicht hergestellt werden. Keine Server-Endpunkte gefunden. @4%s@'; 29 'Verbindung konnte nicht hergestellt werden. Applikation-Instanz-Zertifikat wurde nicht gefunden.'; 30 'Verbindung konnte nicht hergestellt werden. Unerwartetes Format des Zertifikats @4%s@.'; 31 'Verbindung konnte nicht hergestellt werden. Unerwartetes Format der Zertifikatsperrliste @4%s@.'; 32 'Verbindung konnte nicht hergestellt werden. Benutzer konnte nicht authentifiziert werden. Ein Verschlüsselungsdetail ist ungültig. @4%s@'; 34 'Verbindung konnte nicht hergestellt werden. - Der konfigurierte nicht-transparente Redundanzmodus @4%s@ wird nicht unterstützt.'; 101 'Variablen: Adresse @6%s@ existiert nicht auf dem Server.'; 103 'Variablen: Auf Adresse @6%s@ kann nicht zugegriffen werden.'; 104 'Variablen: Erfassungsart wird für Adresse @6%s@ nicht unterstützt.'; 201 'Alarme: Adresse @6%s@ existiert nicht auf dem Server.'; 202 'Alarme: Adresse @6%s@ kann nicht verwendet werden. Der angegebene Bereichsfilter ist kein OPC UA Event notifier.'; 203 'Alarme: Adresse @6%s@ kann nicht verwendet werden. Der angegebene Bereichsfilter existiert nicht auf dem Server.'; 204 'Alarme: Adresse @6%s@ kann nicht verwendet werden, da es sich nicht um einen OPC UA Event type handelt.'; 205 'Alarme: Adresse @6%s@ kann nicht verwendet werden, da der OPC UA Condition type nicht unterstützt wird.'; 206 'Alarme: Adresse @6%s@ kann nicht verwendet werden, da der Event-Typ auf dem Server nicht existiert.'; 207 'Alarme: Erfassungsart kann für Adresse @6%s@ nicht verwendet werden.'; 301 'Adresse @6%s@ kann nicht verwendet werden, da die Versionsnummer fehlt.'; 302 'Adresse @6%s@ kann nicht verwendet werden, da die Versionsnummer ungültig ist.'; 303 'Adresse @6%s@ kann nicht verwendet werden, da die Anzahl der Trennzeichen '$' ungültig ist.'; 304 'Adresse @6%s@ kann nicht verwendet werden, da der Adresstyp ungültig ist.'; 305 'Nicht unterstützte Version @6%s@ der Adresse'; 401 'Nicht erwartete Antwort von OPC UA Server: @6%s@'

text list "SystemTextList_ConfigErrorAlarmTextLibrary_7": 1 'Meldungen: Ungültige Bedingungszeichenfolge für die Alarmanzeige @6%s@.'; 2 'Meldungen: Ungültige Zustandsvariable und Bit für die Alarmanzeige @6%s@.'; 3 'Meldungen: Ungültige Steuervariable und Bit für die Alarmanzeige @6%s@.'

text list "SystemTextList_ConfigErrorAlarmTextLibrary_8": 1 'Archive: Implizites Löschen. Archivvariable-Instanz @6%s@ sollte gelöscht werden. Es existieren aber überladene Elemente.'

text list "SystemTextList_ConfigErrorAlarmTextLibrary_9": 1 ''; 2 'Neustart der Runtime ist erforderlich.'; 3 'Das korrekte Speichermedium muss ausgeworfen und wieder eingelegt werden.'

text list "SystemTextList_ConfigErrorAlarmTextLibrary_10": 1 'CDS-Cache: Cache-Verzeichnis kann nicht erstellt oder erreicht werden: @6%s@'; 2 'LOC-Cache: Cache-Verzeichnis kann nicht erstellt oder erreicht werden: @6%s@'

text list "SystemTextList_RuntimeCollaborationFailureReason_1": 0 'Unbekannter Fehler (@3%s@)'; 1 'Das System läuft nicht oder es besteht ein Netzwerkproblem'; 2 'Auf dem Zielgerät ist Runtime nicht gestartet.'; 3 'Die System-ID stimmt nicht mit der erwarteten System-ID überein @3%s@'; 4 'Der Collaboration-Name stimmt nicht mit dem erwarteten Collaboration-Namen überein '@3%s@''; 5 'Falsches oder unbekanntes Zertifikat'; 6 'Gesperrtes Zertifikat'; 7 'Die Zeitdifferenz ist zu groß.'; 8 'No common supported message version'; 9 'System-ID (@3%s@) existiert bereits'; 10 'Systemname (@3%s@) existiert bereits'; 11 'ID/Name in der lokalen Konfiguration für Runtime Collaboration existiert bereits'

text list "SystemTextList_S7PlusAlarmTextListCollection_1": 4096 'Verbindungen: Verbindung zur PLC @5%s@ getrennt'; 4097 'Verbindungen: Verbindung zum HMI-Gerät @5%s@ getrennt'; 4098 'Verbindungen: Maximale Anzahl von verfügbaren Verbindungen ist überschritten - @5%s@'; 4099 'Nicht genügend Ressourcen auf der PLC verfügbar - @5%s@'; 4100 'Legitimierung fehlgeschlagen, falsches oder fehlendes Passwort - @5%s@'; 4101 'Verbindungsanfrage zum Öffnen der Verbindung fehlgeschlagen - @5%s@'; 4102 'Verbindung: Verbindung zur PLC @5%s@ konnte nicht hergestellt werden'; 4103 'Verbindungsanfrage zum Öffnen der Verbindung konnte nicht gesendet werden'; 4104 'Allgemeiner Zertifikatsfehler für PLC - @5%s@'; 4105 'Das PLC-Zertifikat ist abgelaufen für - @5%s@'; 4106 'PLC Certificate is revoked for - @5%s@'; 4107 'PLC Certificate is untrusted, manual trust is possible for - @5%s@'; 4108 'PLC Certificate is untrusted, manual trust is impossible for - @5%s@'

text list "SystemTextList_AllenBradleyEIPAlarmTextListCollection_7": 4096 'Verbindung PLC-seitig verloren - @5%s@'; 4097 'Verbindung HMI-seitig verloren - @5%s@'; 4098 'Maximale Anzahl von Verbindungen überschritten - @5%s@'; 4099 'Nicht genügend Resourcen auf der PLC verfügbar - @5%s@'; 4100 'Legitimierung fehlgeschlagen, falsches oder fehlendes Passwort - @5%s@'; 4101 'Verbindungsanfrage zum Öffnen der Verbindung fehlgeschlagen - @5%s@'; 4102 'Öffnen der Verbindung fehlgeschlagen - @5%s@'; 4103 'Verbindungsanfrage zum Öffnen der Verbindung konnte nicht gesendet werden'; 4104 'Root Zertifikat ist abgelaufen für - @5%s@'; 4105 'PLC Zertifikat ist ungülzig für - @5%s@'

text list "SystemTextList_OmronEIPAlarmTextListCollection_6": 4096 'Verbindung PLC-seitig verloren - @5%s@'; 4097 'Verbindung HMI-seitig verloren - @5%s@'; 4098 'Maximale Anzahl von Verbindungen überschritten - @5%s@'; 4099 'Nicht genügend Resourcen auf der PLC verfügbar - @5%s@'; 4100 'Legitimierung fehlgeschlagen, falsches oder fehlendes Passwort - @5%s@'; 4101 'Verbindungsanfrage zum Öffnen der Verbindung fehlgeschlagen - @5%s@'; 4102 'Öffnen der Verbindung fehlgeschlagen - @5%s@'; 4103 'Verbindungsanfrage zum Öffnen der Verbindung konnte nicht gesendet werden'; 4104 'Root Zertifikat ist abgelaufen für - @5%s@'; 4105 'PLC Zertifikat ist ungülzig für - @5%s@'

text list "SystemTextList_StdModbusTCPAlarmTextListCollection_5": 4096 'Verbindungen: Verbindung zur PLC @5%s@ getrennt'; 4097 'Verbindungen: Verbindung zum HMI-Gerät @5%s@ getrennt'; 4098 'Verbindungen: Maximale Anzahl von verfügbaren Verbindungen ist überschritten - @5%s@'; 4099 'Nicht genügend Ressourcen auf der PLC verfügbar - @5%s@'; 4100 'Legitimierung fehlgeschlagen, falsches oder fehlendes Passwort - @5%s@'; 4101 'Verbindungsanfrage zum Öffnen der Verbindung fehlgeschlagen - @5%s@'; 4102 'Verbindung: Verbindung zur PLC @5%s@ konnte nicht hergestellt werden'; 4103 'Verbindungsanfrage zum Öffnen der Verbindung konnte nicht gesendet werden'; 4104 'Allgemeiner Zertifikatsfehler für PLC - @5%s@'; 4105 'Das PLC-Zertifikat ist abgelaufen für - @5%s@'; 4106 'Das PLC-Zertifikat ist gesperrt für - @5%s@'; 4107 'Das PLC-Zertifikat ist nicht vertrauenswürdig. Manuelles Vertrauen ist möglich für - @5%s@'; 4108 'Das PLC-Zertifikat ist nicht vertrauenswürdig. Manuelles Vertrauen ist nicht möglich für - @5%s@'

text list "SystemTextList_MitsubishiMCAlarmTextListCollection_4": 4096 'Verbindung PLC-seitig verloren - @5%s@'; 4097 'Verbindung HMI-seitig verloren - @5%s@'; 4098 'Maximale Anzahl von Verbindungen überschritten - @5%s@'; 4099 'Nicht genügend Resourcen auf der PLC verfügbar - @5%s@'; 4100 'Legitimierung fehlgeschlagen, falsches oder fehlendes Passwort - @5%s@'; 4101 'Verbindungsanfrage zum Öffnen der Verbindung fehlgeschlagen - @5%s@'; 4102 'Öffnen der Verbindung fehlgeschlagen - @5%s@'; 4103 'Verbindungsanfrage zum Öffnen der Verbindung konnte nicht gesendet werden'; 4104 'Root Zertifikat ist abgelaufen für - @5%s@'; 4105 'PLC Zertifikat ist ungülzig für - @5%s@'

text list "SystemTextList_MitsubishiiQAlarmTextListCollection_3": 4096 'Verbindung PLC-seitig verloren - @5%s@'; 4097 'Verbindung HMI-seitig verloren - @5%s@'; 4098 'Maximale Anzahl von Verbindungen überschritten - @5%s@'; 4099 'Nicht genügend Resourcen auf der PLC verfügbar - @5%s@'; 4100 'Legitimierung fehlgeschlagen, falsches oder fehlendes Passwort - @5%s@'; 4101 'Verbindungsanfrage zum Öffnen der Verbindung fehlgeschlagen - @5%s@'; 4102 'Öffnen der Verbindung fehlgeschlagen - @5%s@'; 4103 'Verbindungsanfrage zum Öffnen der Verbindung konnte nicht gesendet werden'; 4104 'Root Zertifikat ist abgelaufen für - @5%s@'; 4105 'PLC Zertifikat ist ungülzig für - @5%s@'

text list "SystemTextList_StdModbusRTUAlarmTextListCollection_8": 4096 'Verbindungen: Verbindung zur PLC @5%s@ getrennt'; 4097 'Verbindungen: Verbindung zum HMI-Gerät @5%s@ getrennt'; 4098 'Verbindungen: Maximale Anzahl von verfügbaren Verbindungen ist überschritten - @5%s@'; 4099 'Nicht genügend Ressourcen auf der PLC verfügbar - @5%s@'; 4100 'Legitimierung fehlgeschlagen, falsches oder fehlendes Passwort - @5%s@'; 4101 'Verbindungsanfrage zum Öffnen der Verbindung fehlgeschlagen - @5%s@'; 4102 'Verbindung: Verbindung zur PLC @5%s@ konnte nicht hergestellt werden'; 4103 'Verbindungsanfrage zum Öffnen der Verbindung konnte nicht gesendet werden'; 4104 'Allgemeiner Zertifikatsfehler für PLC - @5%s@'; 4105 'Das PLC-Zertifikat ist abgelaufen für - @5%s@'; 4106 'Das PLC-Zertifikat ist gesperrt für - @5%s@'; 4107 'Das PLC-Zertifikat ist nicht vertrauenswürdig. Manuelles Vertrauen ist möglich für - @5%s@'; 4108 'Das PLC-Zertifikat ist nicht vertrauenswürdig. Manuelles Vertrauen ist nicht möglich für - @5%s@'

graphic list "Grafikliste_1": 0..1 'robotino'; 2..3 'docking2x'; 4..5 'lamptower'; 6..7 'saftey'; 8..9 'robotino-navigation.2'; 10..11 'robotino-carrierBelt'
*)